REGION Network 12
   RUNG wire#powerrail
      Sub(in1 := "EMS".Zone[#Zone].CarrierZnStatus[#PrevZonePos].Position, in2 := "EMS".Zone[#Zone].CarrierSpacing, out => #NextStopPosition)
   END_RUNG
   // the same network as SCL:
   #NextStopPosition := "EMS".Zone[#Zone].CarrierZnStatus[#PrevZonePos].Position - "EMS".Zone[#Zone].CarrierSpacing;
END_REGION

REGION Network 13
   RUNG wire#powerrail
      Sub(in1 := #TrafficCopCarrierZnBuffer[#ZonePos].CommandPos, in2 := "EMS".CoarsePositionDecelOffset, out => #TrafficCopCarrierZnBuffer[#ZonePos].DecelPosition)
   END_RUNG
   // the same network as SCL:
   #TrafficCopCarrierZnBuffer[#ZonePos].DecelPosition := #TrafficCopCarrierZnBuffer[#ZonePos].CommandPos - "EMS".CoarsePositionDecelOffset;
END_REGION

REGION Network 14
   RUNG wire#powerrail
      Contact( "EMS".Carrier[#CarNumZnPos].SDC_IN.AutoMode )
      I_Contact( #TrafficCopCarrierZnBuffer[#ZonePos].AtCommandPos )
      { S7_Templates := "SrcType := DInt" } GT_Contact(in1 := "EMS".Zone[#Zone].CarrierZnStatus[#ZonePos].Position, in2 := #TrafficCopCarrierZnBuffer[#ZonePos].DecelPosition)
      Move(in := "EMS".CoarseDecelSpeed, out1 => #DriveCmdSpeed)
   END_RUNG
   // the same network as SCL:
   IF "EMS".Carrier[#CarNumZnPos].SDC_IN.AutoMode AND NOT #TrafficCopCarrierZnBuffer[#ZonePos].AtCommandPos AND ("EMS".Zone[#Zone].CarrierZnStatus[#ZonePos].Position > #TrafficCopCarrierZnBuffer[#ZonePos].DecelPosition) THEN
       #DriveCmdSpeed := "EMS".CoarseDecelSpeed;
   END_IF;
END_REGION

REGION Network 15
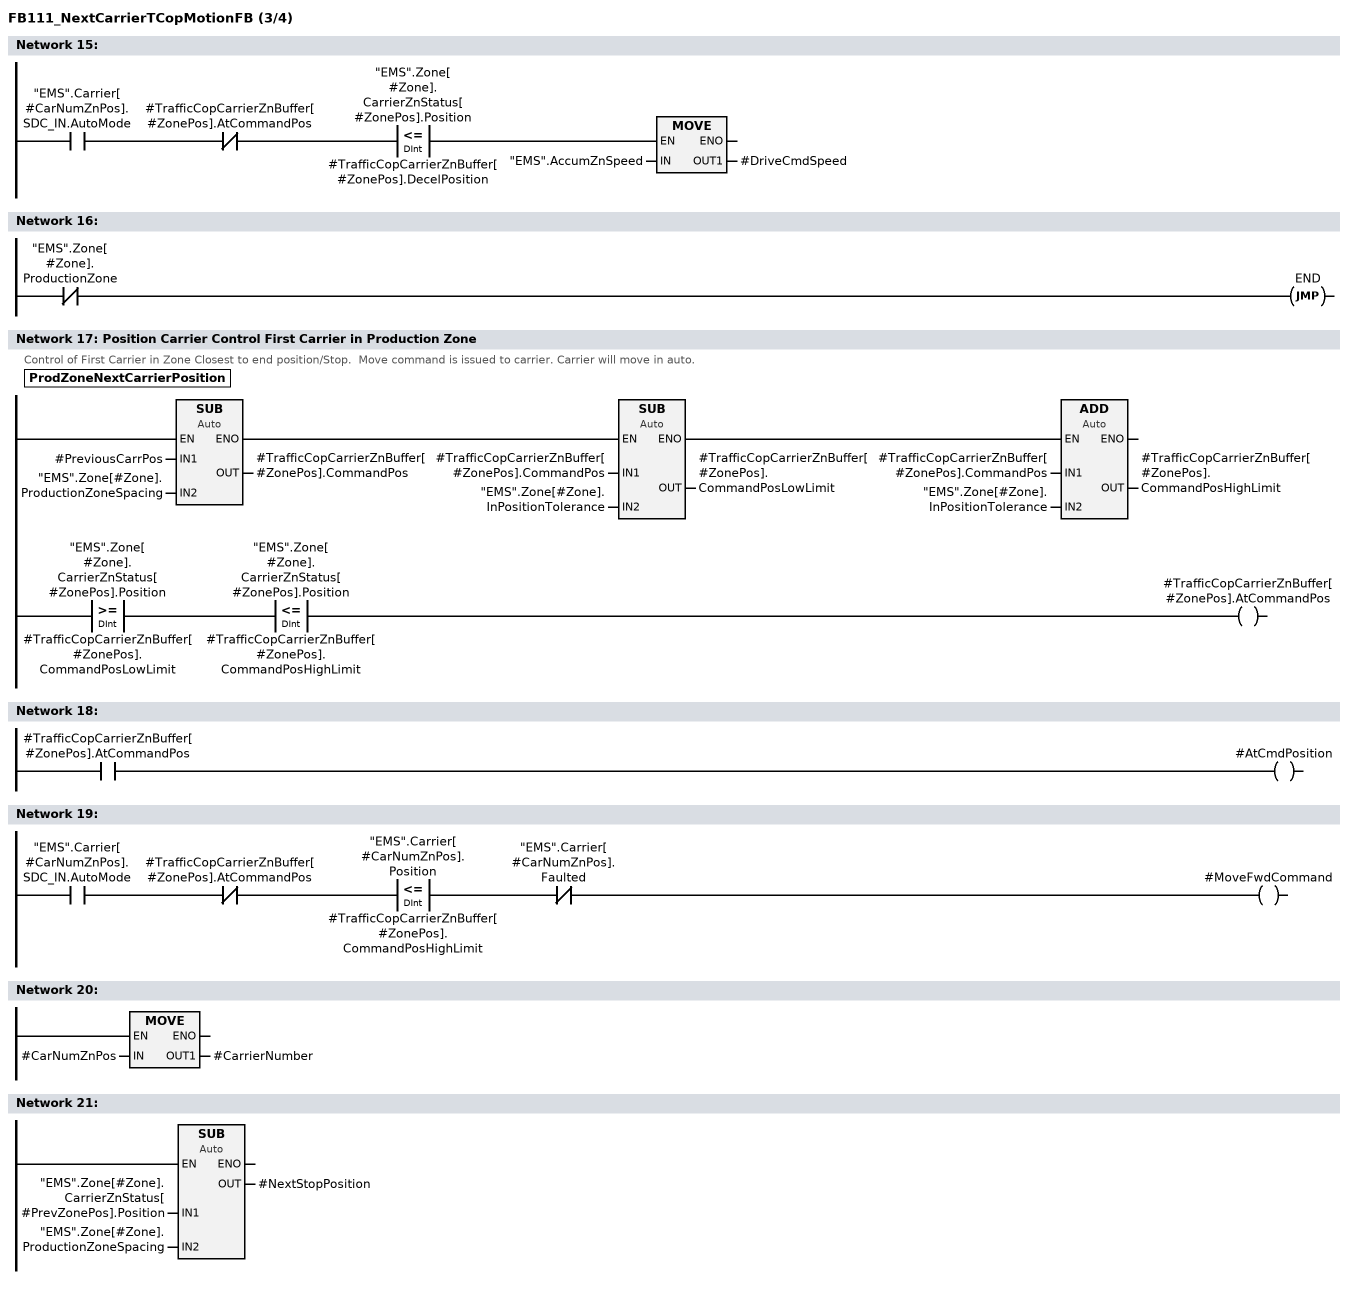
   RUNG wire#powerrail
      Contact( "EMS".Carrier[#CarNumZnPos].SDC_IN.AutoMode )
      I_Contact( #TrafficCopCarrierZnBuffer[#ZonePos].AtCommandPos )
      { S7_Templates := "SrcType := DInt" } LE_Contact(in1 := "EMS".Zone[#Zone].CarrierZnStatus[#ZonePos].Position, in2 := #TrafficCopCarrierZnBuffer[#ZonePos].DecelPosition)
      Move(in := "EMS".AccumZnSpeed, out1 => #DriveCmdSpeed)
   END_RUNG
   // the same network as SCL:
   IF "EMS".Carrier[#CarNumZnPos].SDC_IN.AutoMode AND NOT #TrafficCopCarrierZnBuffer[#ZonePos].AtCommandPos AND ("EMS".Zone[#Zone].CarrierZnStatus[#ZonePos].Position <= #TrafficCopCarrierZnBuffer[#ZonePos].DecelPosition) THEN
       #DriveCmdSpeed := "EMS".AccumZnSpeed;
   END_IF;
END_REGION

REGION Network 16
   RUNG wire#powerrail
      I_Contact( "EMS".Zone[#Zone].ProductionZone )
      JumpCoil( END )
   END_RUNG
   // the same network as SCL:
   IF NOT "EMS".Zone[#Zone].ProductionZone THEN GOTO END; END_IF;
END_REGION

REGION Network 17: Position Carrier Control First Carrier in Production Zone
   // Control of First Carrier in Zone Closest to end position/Stop.  Move command is issued to carrier. Carrier will move in auto.
   Label( ProdZoneNextCarrierPosition )
   RUNG wire#powerrail
      Sub(in1 := #PreviousCarrPos, in2 := "EMS".Zone[#Zone].ProductionZoneSpacing, out => #TrafficCopCarrierZnBuffer[#ZonePos].CommandPos)
      Sub(in1 := #TrafficCopCarrierZnBuffer[#ZonePos].CommandPos, in2 := "EMS".Zone[#Zone].InPositionTolerance, out => #TrafficCopCarrierZnBuffer[#ZonePos].CommandPosLowLimit)
      Add(in1 := #TrafficCopCarrierZnBuffer[#ZonePos].CommandPos, in2 := "EMS".Zone[#Zone].InPositionTolerance, out => #TrafficCopCarrierZnBuffer[#ZonePos].CommandPosHighLimit)
   END_RUNG
   RUNG wire#powerrail
      { S7_Templates := "SrcType := DInt" } GE_Contact(in1 := "EMS".Zone[#Zone].CarrierZnStatus[#ZonePos].Position, in2 := #TrafficCopCarrierZnBuffer[#ZonePos].CommandPosLowLimit)
      { S7_Templates := "SrcType := DInt" } LE_Contact(in1 := "EMS".Zone[#Zone].CarrierZnStatus[#ZonePos].Position, in2 := #TrafficCopCarrierZnBuffer[#ZonePos].CommandPosHighLimit)
      Coil( #TrafficCopCarrierZnBuffer[#ZonePos].AtCommandPos )
   END_RUNG
   // the same network as SCL:
   ProdZoneNextCarrierPosition:
   #TrafficCopCarrierZnBuffer[#ZonePos].CommandPos := #PreviousCarrPos - "EMS".Zone[#Zone].ProductionZoneSpacing;
   #TrafficCopCarrierZnBuffer[#ZonePos].CommandPosLowLimit := #TrafficCopCarrierZnBuffer[#ZonePos].CommandPos - "EMS".Zone[#Zone].InPositionTolerance;
   #TrafficCopCarrierZnBuffer[#ZonePos].CommandPosHighLimit := #TrafficCopCarrierZnBuffer[#ZonePos].CommandPos + "EMS".Zone[#Zone].InPositionTolerance;
   #TrafficCopCarrierZnBuffer[#ZonePos].AtCommandPos := ("EMS".Zone[#Zone].CarrierZnStatus[#ZonePos].Position >= #TrafficCopCarrierZnBuffer[#ZonePos].CommandPosLowLimit) AND ("EMS".Zone[#Zone].CarrierZnStatus[#ZonePos].Position <= #TrafficCopCarrierZnBuffer[#ZonePos].CommandPosHighLimit);
END_REGION

REGION Network 18
   RUNG wire#powerrail
      Contact( #TrafficCopCarrierZnBuffer[#ZonePos].AtCommandPos )
      Coil( #AtCmdPosition )
   END_RUNG
   // the same network as SCL:
   #AtCmdPosition := #TrafficCopCarrierZnBuffer[#ZonePos].AtCommandPos;
END_REGION

REGION Network 19
   RUNG wire#powerrail
      Contact( "EMS".Carrier[#CarNumZnPos].SDC_IN.AutoMode )
      I_Contact( #TrafficCopCarrierZnBuffer[#ZonePos].AtCommandPos )
      { S7_Templates := "SrcType := DInt" } LE_Contact(in1 := "EMS".Carrier[#CarNumZnPos].Position, in2 := #TrafficCopCarrierZnBuffer[#ZonePos].CommandPosHighLimit)
      I_Contact( "EMS".Carrier[#CarNumZnPos].Faulted )
      Coil( #MoveFwdCommand )
   END_RUNG
   // the same network as SCL:
   #MoveFwdCommand := "EMS".Carrier[#CarNumZnPos].SDC_IN.AutoMode AND NOT #TrafficCopCarrierZnBuffer[#ZonePos].AtCommandPos AND ("EMS".Carrier[#CarNumZnPos].Position <= #TrafficCopCarrierZnBuffer[#ZonePos].CommandPosHighLimit) AND NOT "EMS".Carrier[#CarNumZnPos].Faulted;
END_REGION

REGION Network 20
   RUNG wire#powerrail
      Move(in := #CarNumZnPos, out1 => #CarrierNumber)
   END_RUNG
   // the same network as SCL:
   #CarrierNumber := #CarNumZnPos;
END_REGION

REGION Network 21
   RUNG wire#powerrail
      Sub(in1 := "EMS".Zone[#Zone].CarrierZnStatus[#PrevZonePos].Position, in2 := "EMS".Zone[#Zone].ProductionZoneSpacing, out => #NextStopPosition)
   END_RUNG
   // the same network as SCL:
   #NextStopPosition := "EMS".Zone[#Zone].CarrierZnStatus[#PrevZonePos].Position - "EMS".Zone[#Zone].ProductionZoneSpacing;
END_REGION

REGION Network 22
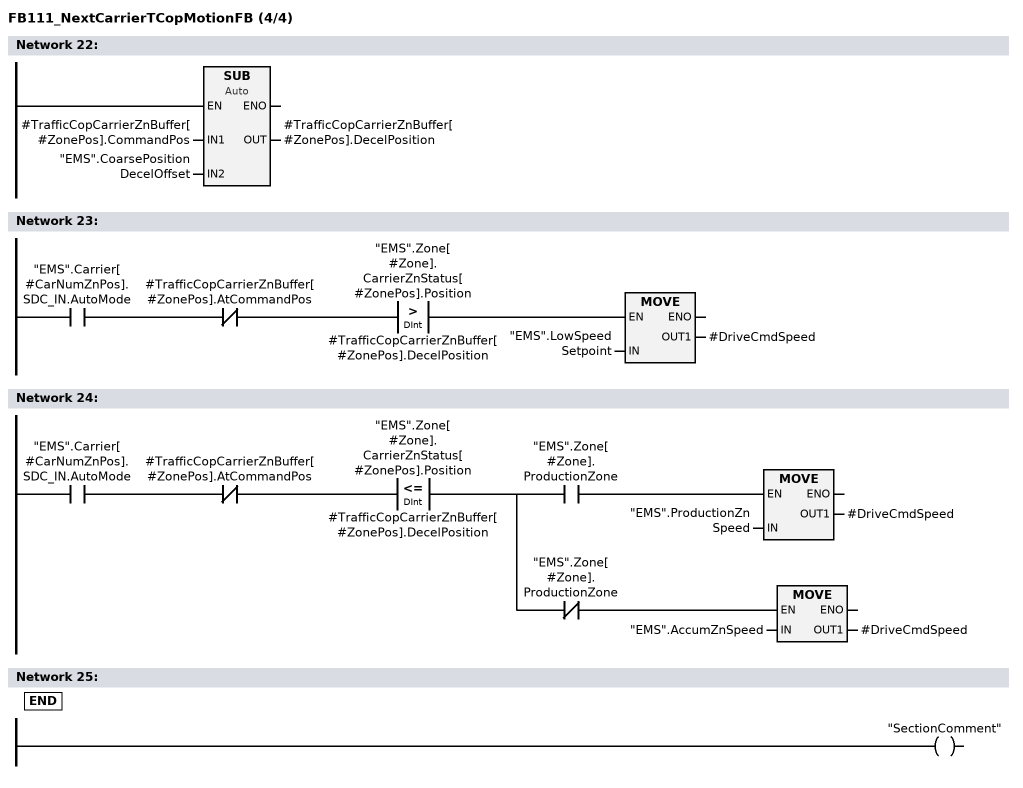
   RUNG wire#powerrail
      Sub(in1 := #TrafficCopCarrierZnBuffer[#ZonePos].CommandPos, in2 := "EMS".CoarsePositionDecelOffset, out => #TrafficCopCarrierZnBuffer[#ZonePos].DecelPosition)
   END_RUNG
   // the same network as SCL:
   #TrafficCopCarrierZnBuffer[#ZonePos].DecelPosition := #TrafficCopCarrierZnBuffer[#ZonePos].CommandPos - "EMS".CoarsePositionDecelOffset;
END_REGION

REGION Network 23
   RUNG wire#powerrail
      Contact( "EMS".Carrier[#CarNumZnPos].SDC_IN.AutoMode )
      I_Contact( #TrafficCopCarrierZnBuffer[#ZonePos].AtCommandPos )
      { S7_Templates := "SrcType := DInt" } GT_Contact(in1 := "EMS".Zone[#Zone].CarrierZnStatus[#ZonePos].Position, in2 := #TrafficCopCarrierZnBuffer[#ZonePos].DecelPosition)
      Move(in := "EMS".LowSpeedSetpoint, out1 => #DriveCmdSpeed)
   END_RUNG
   // the same network as SCL:
   IF "EMS".Carrier[#CarNumZnPos].SDC_IN.AutoMode AND NOT #TrafficCopCarrierZnBuffer[#ZonePos].AtCommandPos AND ("EMS".Zone[#Zone].CarrierZnStatus[#ZonePos].Position > #TrafficCopCarrierZnBuffer[#ZonePos].DecelPosition) THEN
       #DriveCmdSpeed := "EMS".LowSpeedSetpoint;
   END_IF;
END_REGION

REGION Network 24
   RUNG wire#powerrail
      Contact( "EMS".Carrier[#CarNumZnPos].SDC_IN.AutoMode )
      I_Contact( #TrafficCopCarrierZnBuffer[#ZonePos].AtCommandPos )
      { S7_Templates := "SrcType := DInt" } LE_Contact(in1 := "EMS".Zone[#Zone].CarrierZnStatus[#ZonePos].Position, in2 := #TrafficCopCarrierZnBuffer[#ZonePos].DecelPosition)
      wire#w1
      Contact( "EMS".Zone[#Zone].ProductionZone )
      Move(in := "EMS".ProductionZnSpeed, out1 => #DriveCmdSpeed)
   END_RUNG
   RUNG wire#w1
      I_Contact( "EMS".Zone[#Zone].ProductionZone )
      Move(in := "EMS".AccumZnSpeed, out1 => #DriveCmdSpeed)
   END_RUNG
   // the same network as SCL:
   #_w1 := "EMS".Carrier[#CarNumZnPos].SDC_IN.AutoMode AND NOT #TrafficCopCarrierZnBuffer[#ZonePos].AtCommandPos AND ("EMS".Zone[#Zone].CarrierZnStatus[#ZonePos].Position <= #TrafficCopCarrierZnBuffer[#ZonePos].DecelPosition);
   IF #_w1 AND "EMS".Zone[#Zone].ProductionZone THEN #DriveCmdSpeed := "EMS".ProductionZnSpeed; END_IF;
   IF #_w1 AND NOT "EMS".Zone[#Zone].ProductionZone THEN #DriveCmdSpeed := "EMS".AccumZnSpeed; END_IF;
END_REGION

REGION Network 25
   Label( END )
   RUNG wire#powerrail
      Coil( "SectionComment" )
   END_RUNG
   // the same network as SCL:
   END:
   "SectionComment" := TRUE;
END_REGION
END_FUNCTION_BLOCK

FUNCTION_BLOCK "FB112_Carrier"   // FB112, LAD
{ S7_Optimized_Access := 'TRUE' }
VERSION : 0.1
   VAR_INPUT
      Carrier : Int;
      EMS : "UDT_System";
      MoveFwd : Bool;
      SpeedSelect : Word;   // Speed Select 1=Slow 2=Normal
      CarrierFindArrayBufferiN : "UDT_Carrier";
      SDC_IN : "UDT_SDC_IN";
      DuplicateCarrierNumIn : Int;
      DuplicateCarrierFound : Bool;
      GapSpacingFault : Bool;
      FaultReset : Bool;
   END_VAR
   VAR_OUTPUT
      Zone : Int;
      Area : String[2];
      AreaInt : Int;
      ZonePos : Word;
      CarrierPositionEcho : DWord;
      CarrierNumberEcho : Word;
      DuplicateCarrierNumEcho : Word;
      CarrierNextStopPosEcho : Word;
      Faults : "UDT_SDCOutFaults";
      Faulted : Bool;
   END_VAR
   VAR
      CarrierMoveFwdSetup : Array[0..30] of Bool;
      MotionOffFaultTimer : IEC_TIMER;
      MotionOnFaultTimer : IEC_TIMER;
   END_VAR
   VAR_TEMP
      RetVal : Int;
      srcindex : DInt;
      destindex : DInt;
   END_VAR
BEGIN

REGION Network 1
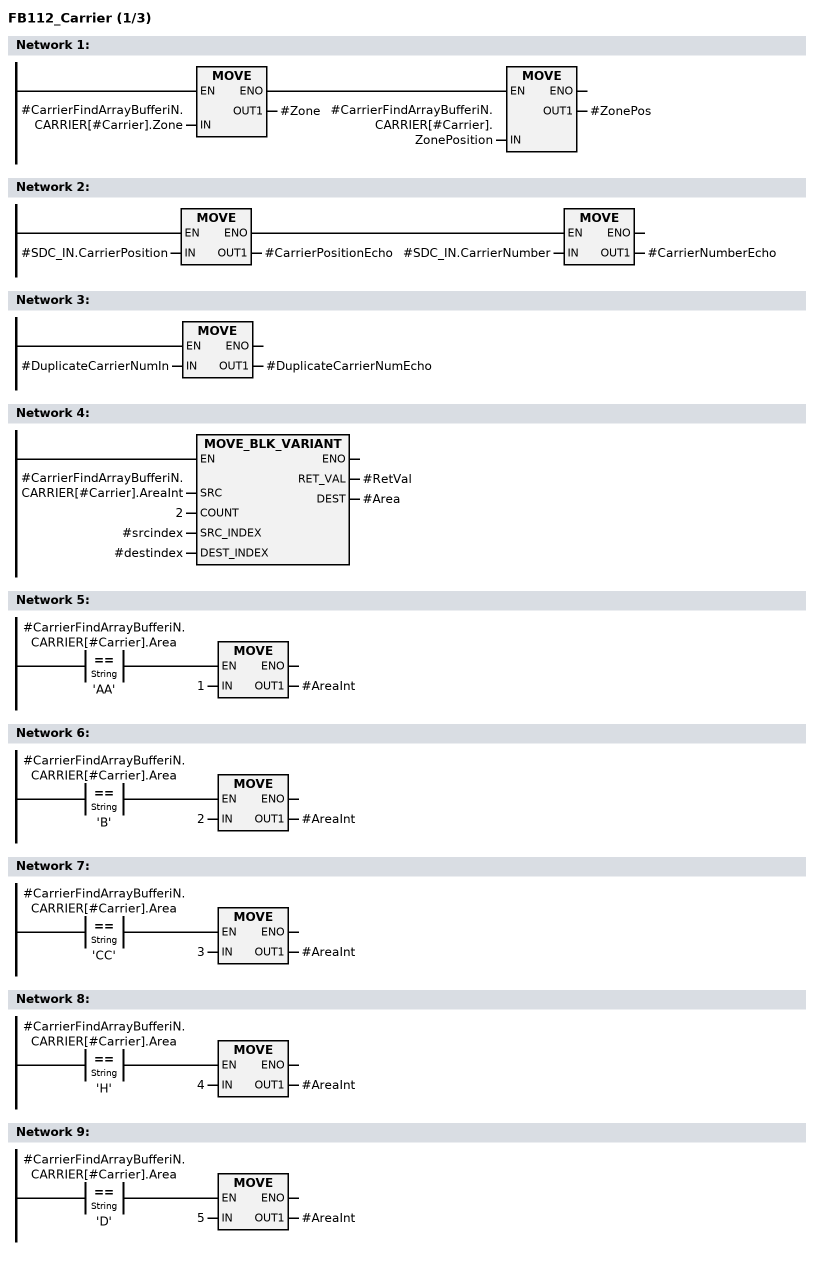
   RUNG wire#powerrail
      Move(in := #CarrierFindArrayBufferiN.CARRIER[#Carrier].Zone, out1 => #Zone)
      Move(in := #CarrierFindArrayBufferiN.CARRIER[#Carrier].ZonePosition, out1 => #ZonePos)
   END_RUNG
   // the same network as SCL:
   #Zone := #CarrierFindArrayBufferiN.CARRIER[#Carrier].Zone;
   #ZonePos := #CarrierFindArrayBufferiN.CARRIER[#Carrier].ZonePosition;
END_REGION

REGION Network 2
   RUNG wire#powerrail
      Move(in := #SDC_IN.CarrierPosition, out1 => #CarrierPositionEcho)
      Move(in := #SDC_IN.CarrierNumber, out1 => #CarrierNumberEcho)
   END_RUNG
   // the same network as SCL:
   #CarrierPositionEcho := #SDC_IN.CarrierPosition;
   #CarrierNumberEcho := #SDC_IN.CarrierNumber;
END_REGION

REGION Network 3
   RUNG wire#powerrail
      Move(in := #DuplicateCarrierNumIn, out1 => #DuplicateCarrierNumEcho)
   END_RUNG
   // the same network as SCL:
   #DuplicateCarrierNumEcho := #DuplicateCarrierNumIn;
END_REGION

REGION Network 4
   #RetVal := MOVE_BLK_VARIANT(SRC := #CarrierFindArrayBufferiN.CARRIER[#Carrier].AreaInt,
                           COUNT := 2,
                           SRC_INDEX := #srcindex,
                           DEST_INDEX := #destindex,
                           DEST => #Area);
END_REGION

REGION Network 5
   RUNG wire#powerrail
      { S7_Templates := "SrcType := String" } EQ_Contact(in1 := #CarrierFindArrayBufferiN.CARRIER[#Carrier].Area, in2 := 'AA')
      Move(in := 1, out1 => #AreaInt)
   END_RUNG
   // the same network as SCL:
   IF #CarrierFindArrayBufferiN.CARRIER[#Carrier].Area = 'AA' THEN #AreaInt := 1; END_IF;
END_REGION

REGION Network 6
   RUNG wire#powerrail
      { S7_Templates := "SrcType := String" } EQ_Contact(in1 := #CarrierFindArrayBufferiN.CARRIER[#Carrier].Area, in2 := 'B')
      Move(in := 2, out1 => #AreaInt)
   END_RUNG
   // the same network as SCL:
   IF #CarrierFindArrayBufferiN.CARRIER[#Carrier].Area = 'B' THEN #AreaInt := 2; END_IF;
END_REGION

REGION Network 7
   RUNG wire#powerrail
      { S7_Templates := "SrcType := String" } EQ_Contact(in1 := #CarrierFindArrayBufferiN.CARRIER[#Carrier].Area, in2 := 'CC')
      Move(in := 3, out1 => #AreaInt)
   END_RUNG
   // the same network as SCL:
   IF #CarrierFindArrayBufferiN.CARRIER[#Carrier].Area = 'CC' THEN #AreaInt := 3; END_IF;
END_REGION

REGION Network 8
   RUNG wire#powerrail
      { S7_Templates := "SrcType := String" } EQ_Contact(in1 := #CarrierFindArrayBufferiN.CARRIER[#Carrier].Area, in2 := 'H')
      Move(in := 4, out1 => #AreaInt)
   END_RUNG
   // the same network as SCL:
   IF #CarrierFindArrayBufferiN.CARRIER[#Carrier].Area = 'H' THEN #AreaInt := 4; END_IF;
END_REGION

REGION Network 9
   RUNG wire#powerrail
      { S7_Templates := "SrcType := String" } EQ_Contact(in1 := #CarrierFindArrayBufferiN.CARRIER[#Carrier].Area, in2 := 'D')
      Move(in := 5, out1 => #AreaInt)
   END_RUNG
   // the same network as SCL:
   IF #CarrierFindArrayBufferiN.CARRIER[#Carrier].Area = 'D' THEN #AreaInt := 5; END_IF;
END_REGION

REGION Network 10
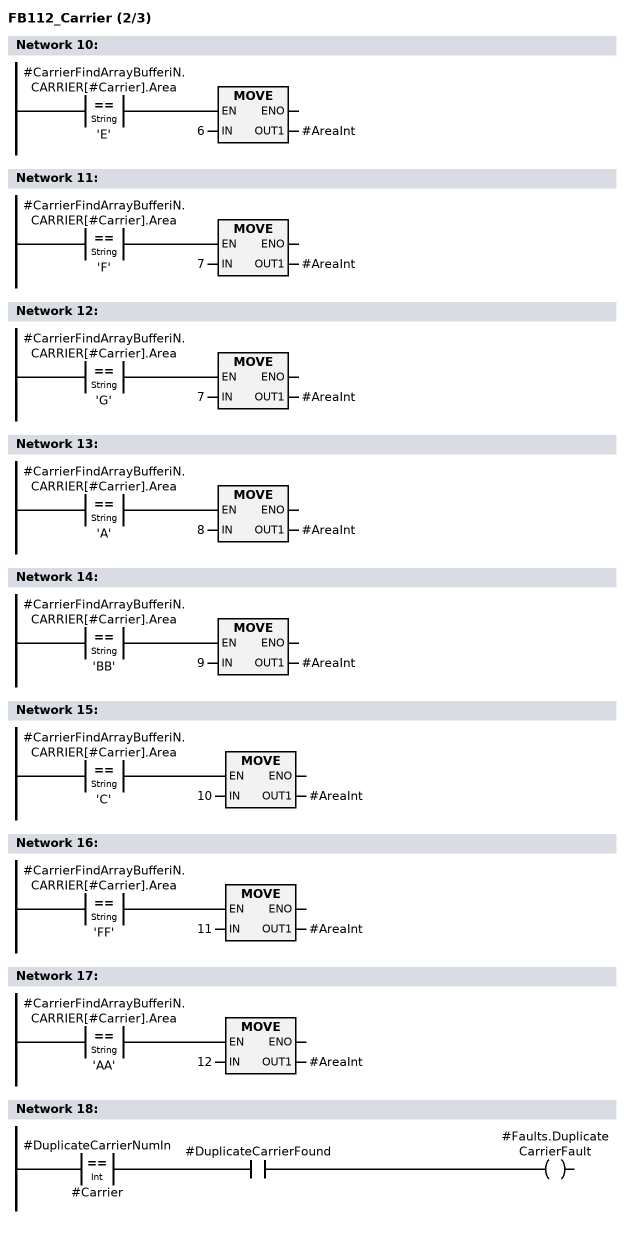
   RUNG wire#powerrail
      { S7_Templates := "SrcType := String" } EQ_Contact(in1 := #CarrierFindArrayBufferiN.CARRIER[#Carrier].Area, in2 := 'E')
      Move(in := 6, out1 => #AreaInt)
   END_RUNG
   // the same network as SCL:
   IF #CarrierFindArrayBufferiN.CARRIER[#Carrier].Area = 'E' THEN #AreaInt := 6; END_IF;
END_REGION

REGION Network 11
   RUNG wire#powerrail
      { S7_Templates := "SrcType := String" } EQ_Contact(in1 := #CarrierFindArrayBufferiN.CARRIER[#Carrier].Area, in2 := 'F')
      Move(in := 7, out1 => #AreaInt)
   END_RUNG
   // the same network as SCL:
   IF #CarrierFindArrayBufferiN.CARRIER[#Carrier].Area = 'F' THEN #AreaInt := 7; END_IF;
END_REGION

REGION Network 12
   RUNG wire#powerrail
      { S7_Templates := "SrcType := String" } EQ_Contact(in1 := #CarrierFindArrayBufferiN.CARRIER[#Carrier].Area, in2 := 'G')
      Move(in := 7, out1 => #AreaInt)
   END_RUNG
   // the same network as SCL:
   IF #CarrierFindArrayBufferiN.CARRIER[#Carrier].Area = 'G' THEN #AreaInt := 7; END_IF;
END_REGION

REGION Network 13
   RUNG wire#powerrail
      { S7_Templates := "SrcType := String" } EQ_Contact(in1 := #CarrierFindArrayBufferiN.CARRIER[#Carrier].Area, in2 := 'A')
      Move(in := 8, out1 => #AreaInt)
   END_RUNG
   // the same network as SCL:
   IF #CarrierFindArrayBufferiN.CARRIER[#Carrier].Area = 'A' THEN #AreaInt := 8; END_IF;
END_REGION

REGION Network 14
   RUNG wire#powerrail
      { S7_Templates := "SrcType := String" } EQ_Contact(in1 := #CarrierFindArrayBufferiN.CARRIER[#Carrier].Area, in2 := 'BB')
      Move(in := 9, out1 => #AreaInt)
   END_RUNG
   // the same network as SCL:
   IF #CarrierFindArrayBufferiN.CARRIER[#Carrier].Area = 'BB' THEN #AreaInt := 9; END_IF;
END_REGION

REGION Network 15
   RUNG wire#powerrail
      { S7_Templates := "SrcType := String" } EQ_Contact(in1 := #CarrierFindArrayBufferiN.CARRIER[#Carrier].Area, in2 := 'C')
      Move(in := 10, out1 => #AreaInt)
   END_RUNG
   // the same network as SCL:
   IF #CarrierFindArrayBufferiN.CARRIER[#Carrier].Area = 'C' THEN #AreaInt := 10; END_IF;
END_REGION

REGION Network 16
   RUNG wire#powerrail
      { S7_Templates := "SrcType := String" } EQ_Contact(in1 := #CarrierFindArrayBufferiN.CARRIER[#Carrier].Area, in2 := 'FF')
      Move(in := 11, out1 => #AreaInt)
   END_RUNG
   // the same network as SCL:
   IF #CarrierFindArrayBufferiN.CARRIER[#Carrier].Area = 'FF' THEN #AreaInt := 11; END_IF;
END_REGION

REGION Network 17
   RUNG wire#powerrail
      { S7_Templates := "SrcType := String" } EQ_Contact(in1 := #CarrierFindArrayBufferiN.CARRIER[#Carrier].Area, in2 := 'AA')
      Move(in := 12, out1 => #AreaInt)
   END_RUNG
   // the same network as SCL:
   IF #CarrierFindArrayBufferiN.CARRIER[#Carrier].Area = 'AA' THEN #AreaInt := 12; END_IF;
END_REGION

REGION Network 18
   RUNG wire#powerrail
      { S7_Templates := "SrcType := Int" } EQ_Contact(in1 := #DuplicateCarrierNumIn, in2 := #Carrier)
      Contact( #DuplicateCarrierFound )
      Coil( #Faults.DuplicateCarrierFault )
   END_RUNG
   // the same network as SCL:
   #Faults.DuplicateCarrierFault := (#DuplicateCarrierNumIn = #Carrier) AND #DuplicateCarrierFound;
END_REGION

REGION Network 19
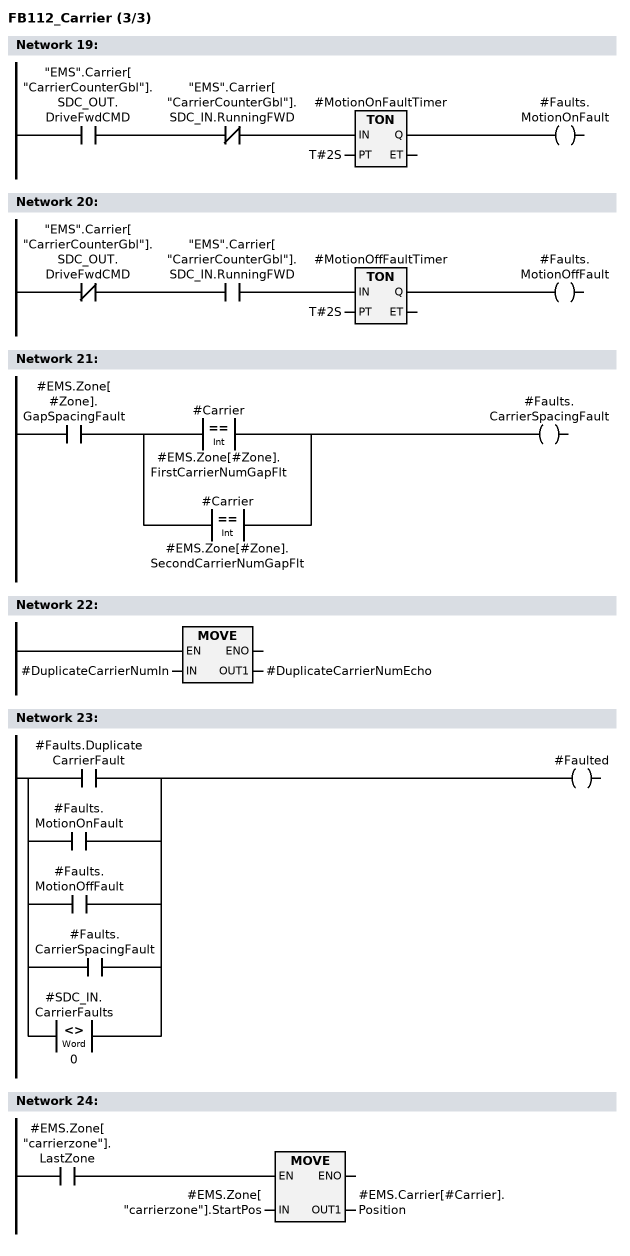
   #MotionOnFaultTimer.TON(IN := "EMS".Carrier["CarrierCounterGbl"].SDC_OUT.DriveFwdCMD AND NOT "EMS".Carrier["CarrierCounterGbl"].SDC_IN.RunningFWD,
                           PT := T#2S);
   #Faults.MotionOnFault := #MotionOnFaultTimer.Q;
END_REGION

REGION Network 20
   #MotionOffFaultTimer.TON(IN := NOT "EMS".Carrier["CarrierCounterGbl"].SDC_OUT.DriveFwdCMD AND "EMS".Carrier["CarrierCounterGbl"].SDC_IN.RunningFWD,
                           PT := T#2S);
   #Faults.MotionOffFault := #MotionOffFaultTimer.Q;
END_REGION

REGION Network 21
   RUNG wire#powerrail
      Contact( #EMS.Zone[#Zone].GapSpacingFault )
      wire#w1
      { S7_Templates := "SrcType := Int" } EQ_Contact(in1 := #Carrier, in2 := #EMS.Zone[#Zone].FirstCarrierNumGapFlt)
      wire#w2
      Coil( #Faults.CarrierSpacingFault )
   END_RUNG
   RUNG wire#w1
      { S7_Templates := "SrcType := Int" } EQ_Contact(in1 := #Carrier, in2 := #EMS.Zone[#Zone].SecondCarrierNumGapFlt)
   END_RUNG wire#w2
   // the same network as SCL:
   #Faults.CarrierSpacingFault := #EMS.Zone[#Zone].GapSpacingFault AND ((#Carrier = #EMS.Zone[#Zone].FirstCarrierNumGapFlt) OR (#Carrier = #EMS.Zone[#Zone].SecondCarrierNumGapFlt));
END_REGION

REGION Network 22
   RUNG wire#powerrail
      Move(in := #DuplicateCarrierNumIn, out1 => #DuplicateCarrierNumEcho)
   END_RUNG
   // the same network as SCL:
   #DuplicateCarrierNumEcho := #DuplicateCarrierNumIn;
END_REGION

REGION Network 23
   RUNG wire#powerrail
      Contact( #Faults.DuplicateCarrierFault )
      wire#w1
      Coil( #Faulted )
   END_RUNG
   RUNG wire#powerrail
      Contact( #Faults.MotionOnFault )
   END_RUNG wire#w1
   RUNG wire#powerrail
      Contact( #Faults.MotionOffFault )
   END_RUNG wire#w1
   RUNG wire#powerrail
      Contact( #Faults.CarrierSpacingFault )
   END_RUNG wire#w1
   RUNG wire#powerrail
      { S7_Templates := "SrcType := Word" } NE_Contact(in1 := #SDC_IN.CarrierFaults, in2 := 0)
   END_RUNG wire#w1
   // the same network as SCL:
   #Faulted := #Faults.DuplicateCarrierFault OR #Faults.MotionOnFault OR #Faults.MotionOffFault OR #Faults.CarrierSpacingFault OR (#SDC_IN.CarrierFaults <> 0);
END_REGION

REGION Network 24
   RUNG wire#powerrail
      Contact( #EMS.Zone["carrierzone"].LastZone )
      Move(in := #EMS.Zone["carrierzone"].StartPos, out1 => #EMS.Carrier[#Carrier].Position)
   END_RUNG
   // the same network as SCL:
   IF #EMS.Zone["carrierzone"].LastZone THEN
       #EMS.Carrier[#Carrier].Position := #EMS.Zone["carrierzone"].StartPos;
   END_IF;
END_REGION
END_FUNCTION_BLOCK

FUNCTION_BLOCK "FB113_CarrierTrafficCop"   // FB113, LAD
{ S7_Optimized_Access := 'TRUE' }
VERSION : 0.1
   VAR_INPUT
      CarrierNumber : Word;
      ZonePos : Word;
   END_VAR
BEGIN
END_FUNCTION_BLOCK

FUNCTION_BLOCK "FB115_FB_Zone"   // FB115, LAD
{ S7_Optimized_Access := 'FALSE' }
VERSION : 0.1
   VAR_INPUT
      Zone : Int;
      Description : String[10];
      LastZone : Bool;
      MaxCarriers : Int;
      StartPos : DWord;
      EndPos : DWord;
      NextZone : Word;   // If Zone numbering is non sequential Next Zone Nu
      PreviousZone : Word;   // If Zone numbering is non sequential Previous Zone Nu
      SpeedZone : Bool;
      SpeedZoneStart : DWord;
      SpeedZoneEnd : DWord;
      AccumZone : Bool;
      AccumZnSpacing : Word;
      ProductionZone : Bool := false;
      ProductZoneSpacing : Word;
      FinePosStopZone : Bool;
      FineInPosTolerance : Word;
      FinePositionDecelOffset : Word;
      CoarseInPosTolerance : Word;
      CoarsePositionDecelOffset : Word;
      NextCarrierClrHighSpeed : Word;
   END_VAR
   VAR_OUTPUT
      ZoneEcho : Word;
      LastZoneEcho : Bool;
      ZoneFull : Bool;
      ZoneLengthEcho : Word;
      DescriptionEcho : String[10];
      StartPosEcho : DWord;
      EndPosEcho : DWord;
      SpeedZoneEcho : Bool;
      SpeedZoneStartEcho : DWord;
      SpeedZoneEndEcho : DWord;
      AccumZoneEcho : Bool;
      AccumSpacingEcho : Word;
      ProductionZoneEcho : Bool;
      ProdZoneSpacingEcho : Word;
      CarrierInPosToleranceEcho : Word;
      NextCarrierClrHighSpeedEcho : Word;
      MaxCarriersEcho : Word;
      ClearToEnterEcho : Bool;
      ClearZoneStartEcho : Bool;
      ClearZoneEcho : Bool;
      ZoneCarrierStatsArray : Array[0..60] of "UDT_ZoneCarrierStatus";
      FinePosStopZoneEcho : Bool;
      FineInPosToleranceEcho : Word;
      FinePositionDecelEcho : Word;
      CoarsePositionDecelEcho : Word;
      CoarseInPosToleranceEcho : Word;
      PreviosZoneEcho : Word;
      NextZoneEcho : Word;
      CarrierAtStop : Bool;
      CarrierNumAtStop : Word;
      HMIZonePositionsEcho : Array[1..20] of "UDT_HMIZonePositions";
      ClearOfStopPos : DWord;
   END_VAR
   VAR_TEMP
      HMIZonePositions : Array[1..20] of "UDT_HMIZonePositions";
      carrierstatusdn : Bool;
      resettemp : Bool;
      resettemp2 : Bool;
      sortdonetemp : Bool;
      ZonePosSpacing : Word;
      ZoneLengthTemp : UDInt;
   END_VAR
BEGIN

REGION Network 1
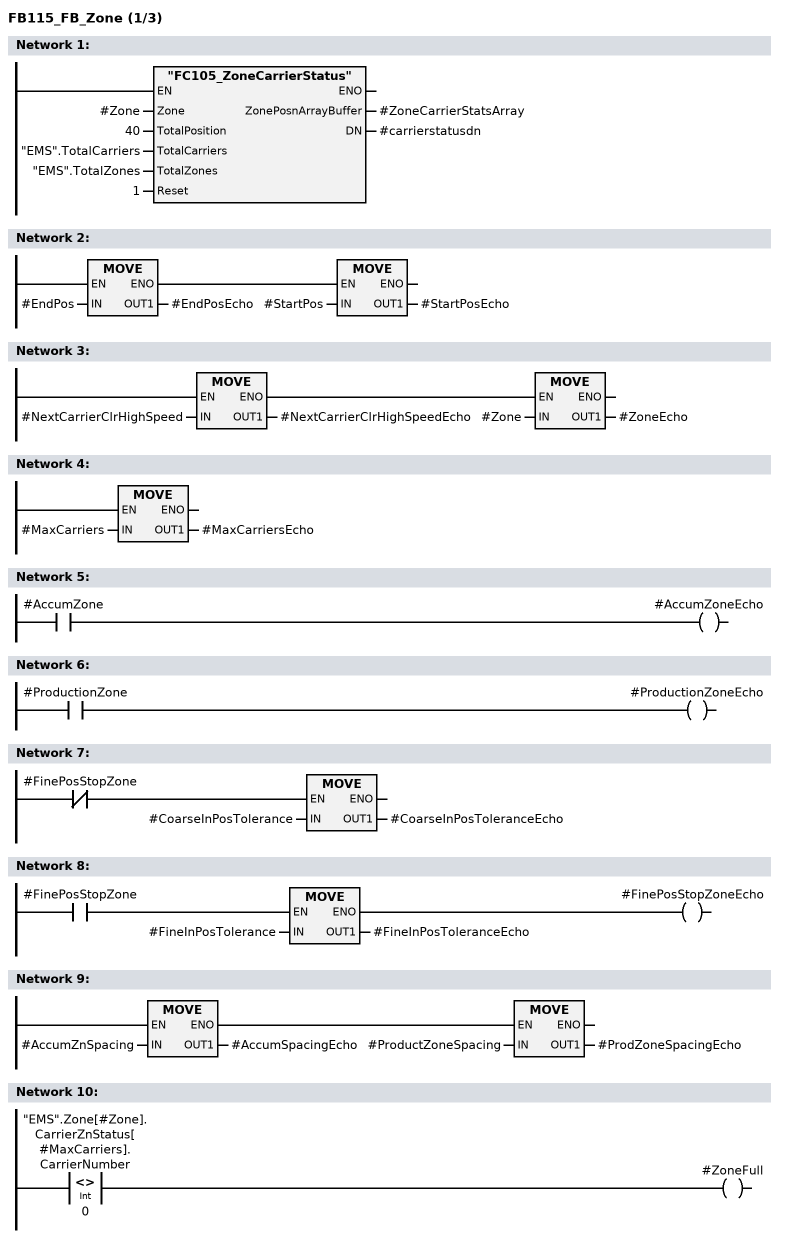
   RUNG wire#powerrail
      "FC105_ZoneCarrierStatus"(Zone := #Zone, TotalPosition := 40, TotalCarriers := "EMS".TotalCarriers, TotalZones := "EMS".TotalZones, Reset := 1, ZonePosnArrayBuffer => #ZoneCarrierStatsArray, DN => #carrierstatusdn)
   END_RUNG
   // the same network as SCL:
   "FC105_ZoneCarrierStatus"(Zone := #Zone,
                           TotalPosition := 40,
                           TotalCarriers := "EMS".TotalCarriers,
                           TotalZones := "EMS".TotalZones,
                           Reset := 1,
                           ZonePosnArrayBuffer => #ZoneCarrierStatsArray,
                           DN => #carrierstatusdn);
END_REGION

REGION Network 2
   RUNG wire#powerrail
      Move(in := #EndPos, out1 => #EndPosEcho)
      Move(in := #StartPos, out1 => #StartPosEcho)
   END_RUNG
   // the same network as SCL:
   #EndPosEcho := #EndPos;
   #StartPosEcho := #StartPos;
END_REGION

REGION Network 3
   RUNG wire#powerrail
      Move(in := #NextCarrierClrHighSpeed, out1 => #NextCarrierClrHighSpeedEcho)
      Move(in := #Zone, out1 => #ZoneEcho)
   END_RUNG
   // the same network as SCL:
   #NextCarrierClrHighSpeedEcho := #NextCarrierClrHighSpeed;
   #ZoneEcho := #Zone;
END_REGION

REGION Network 4
   RUNG wire#powerrail
      Move(in := #MaxCarriers, out1 => #MaxCarriersEcho)
   END_RUNG
   // the same network as SCL:
   #MaxCarriersEcho := #MaxCarriers;
END_REGION

REGION Network 5
   RUNG wire#powerrail
      Contact( #AccumZone )
      Coil( #AccumZoneEcho )
   END_RUNG
   // the same network as SCL:
   #AccumZoneEcho := #AccumZone;
END_REGION

REGION Network 6
   RUNG wire#powerrail
      Contact( #ProductionZone )
      Coil( #ProductionZoneEcho )
   END_RUNG
   // the same network as SCL:
   #ProductionZoneEcho := #ProductionZone;
END_REGION

REGION Network 7
   RUNG wire#powerrail
      I_Contact( #FinePosStopZone )
      Move(in := #CoarseInPosTolerance, out1 => #CoarseInPosToleranceEcho)
   END_RUNG
   // the same network as SCL:
   IF NOT #FinePosStopZone THEN #CoarseInPosToleranceEcho := #CoarseInPosTolerance; END_IF;
END_REGION

REGION Network 8
   RUNG wire#powerrail
      Contact( #FinePosStopZone )
      Move(in := #FineInPosTolerance, out1 => #FineInPosToleranceEcho)
      Coil( #FinePosStopZoneEcho )
   END_RUNG
   // the same network as SCL:
   IF #FinePosStopZone THEN #FineInPosToleranceEcho := #FineInPosTolerance; END_IF;
   #FinePosStopZoneEcho := #FinePosStopZone;
END_REGION

